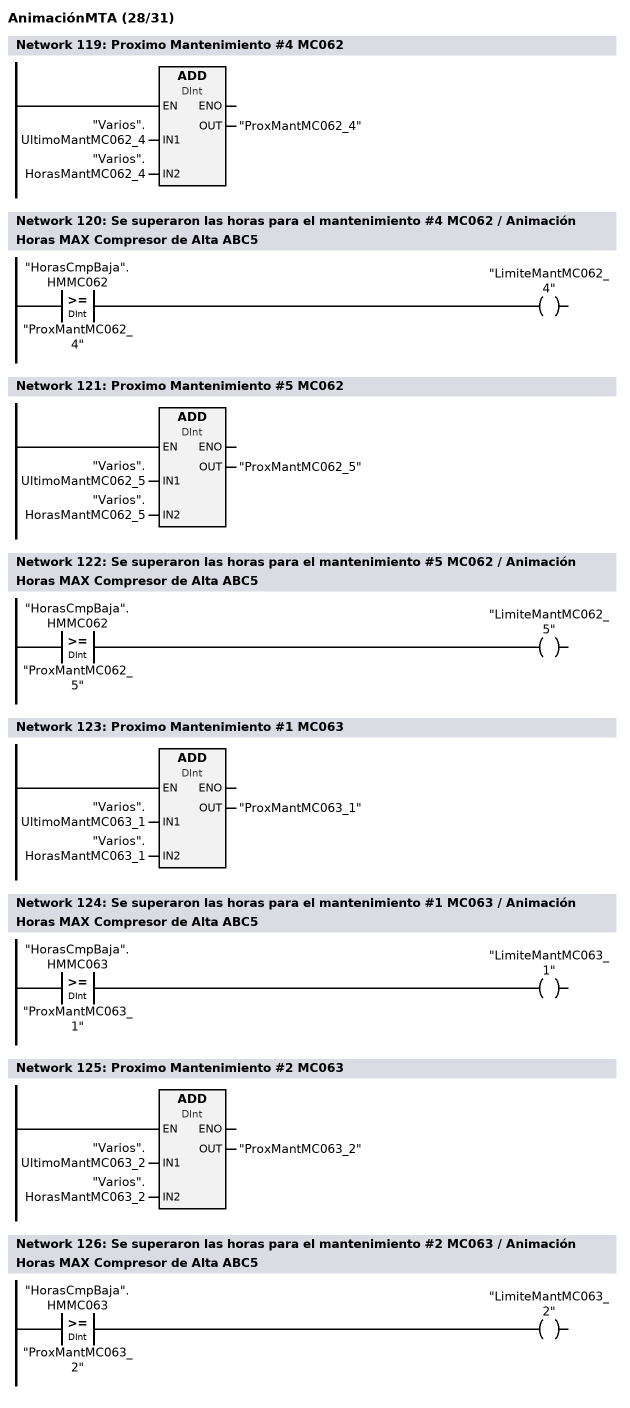
   RUNG wire#powerrail
      { S7_Templates := "SrcType := DInt"; S7_GenerateENO := "TRUE" } Add(in1 := "Varios".UltimoMantMC062_4, in2 := "Varios".HorasMantMC062_4, out => "ProxMantMC062_4")
   END_RUNG
   // the same network as SCL:
   "ProxMantMC062_4" := "Varios".UltimoMantMC062_4 + "Varios".HorasMantMC062_4;
END_REGION

REGION Network 120: Se superaron las horas para el mantenimiento #4 MC062 / Animación Horas MAX Compresor de Alta ABC5
   RUNG wire#powerrail
      { S7_Templates := "SrcType := DInt" } GE_Contact(in1 := "HorasCmpBaja".HMMC062, in2 := "ProxMantMC062_4")
      Coil( "LimiteMantMC062_4" )
   END_RUNG
   // the same network as SCL:
   "LimiteMantMC062_4" := "HorasCmpBaja".HMMC062 >= "ProxMantMC062_4";
END_REGION

REGION Network 121: Proximo Mantenimiento #5 MC062
   RUNG wire#powerrail
      { S7_Templates := "SrcType := DInt"; S7_GenerateENO := "TRUE" } Add(in1 := "Varios".UltimoMantMC062_5, in2 := "Varios".HorasMantMC062_5, out => "ProxMantMC062_5")
   END_RUNG
   // the same network as SCL:
   "ProxMantMC062_5" := "Varios".UltimoMantMC062_5 + "Varios".HorasMantMC062_5;
END_REGION

REGION Network 122: Se superaron las horas para el mantenimiento #5 MC062 / Animación Horas MAX Compresor de Alta ABC5
   RUNG wire#powerrail
      { S7_Templates := "SrcType := DInt" } GE_Contact(in1 := "HorasCmpBaja".HMMC062, in2 := "ProxMantMC062_5")
      Coil( "LimiteMantMC062_5" )
   END_RUNG
   // the same network as SCL:
   "LimiteMantMC062_5" := "HorasCmpBaja".HMMC062 >= "ProxMantMC062_5";
END_REGION

REGION Network 123: Proximo Mantenimiento #1 MC063
   RUNG wire#powerrail
      { S7_Templates := "SrcType := DInt"; S7_GenerateENO := "TRUE" } Add(in1 := "Varios".UltimoMantMC063_1, in2 := "Varios".HorasMantMC063_1, out => "ProxMantMC063_1")
   END_RUNG
   // the same network as SCL:
   "ProxMantMC063_1" := "Varios".UltimoMantMC063_1 + "Varios".HorasMantMC063_1;
END_REGION

REGION Network 124: Se superaron las horas para el mantenimiento #1 MC063 / Animación Horas MAX Compresor de Alta ABC5
   RUNG wire#powerrail
      { S7_Templates := "SrcType := DInt" } GE_Contact(in1 := "HorasCmpBaja".HMMC063, in2 := "ProxMantMC063_1")
      Coil( "LimiteMantMC063_1" )
   END_RUNG
   // the same network as SCL:
   "LimiteMantMC063_1" := "HorasCmpBaja".HMMC063 >= "ProxMantMC063_1";
END_REGION

REGION Network 125: Proximo Mantenimiento #2 MC063
   RUNG wire#powerrail
      { S7_Templates := "SrcType := DInt"; S7_GenerateENO := "TRUE" } Add(in1 := "Varios".UltimoMantMC063_2, in2 := "Varios".HorasMantMC063_2, out => "ProxMantMC063_2")
   END_RUNG
   // the same network as SCL:
   "ProxMantMC063_2" := "Varios".UltimoMantMC063_2 + "Varios".HorasMantMC063_2;
END_REGION

REGION Network 126: Se superaron las horas para el mantenimiento #2 MC063 / Animación Horas MAX Compresor de Alta ABC5
   RUNG wire#powerrail
      { S7_Templates := "SrcType := DInt" } GE_Contact(in1 := "HorasCmpBaja".HMMC063, in2 := "ProxMantMC063_2")
      Coil( "LimiteMantMC063_2" )
   END_RUNG
   // the same network as SCL:
   "LimiteMantMC063_2" := "HorasCmpBaja".HMMC063 >= "ProxMantMC063_2";
END_REGION

REGION Network 127: Proximo Mantenimiento #3 MC063
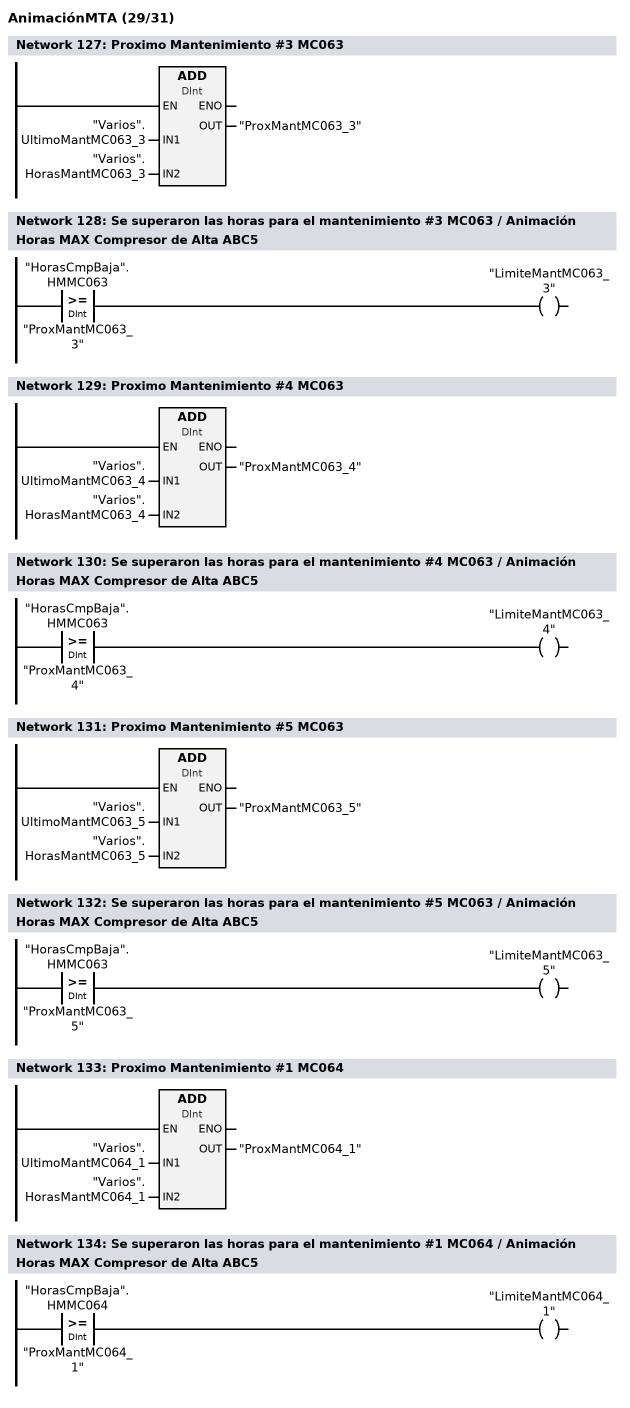
   RUNG wire#powerrail
      { S7_Templates := "SrcType := DInt"; S7_GenerateENO := "TRUE" } Add(in1 := "Varios".UltimoMantMC063_3, in2 := "Varios".HorasMantMC063_3, out => "ProxMantMC063_3")
   END_RUNG
   // the same network as SCL:
   "ProxMantMC063_3" := "Varios".UltimoMantMC063_3 + "Varios".HorasMantMC063_3;
END_REGION

REGION Network 128: Se superaron las horas para el mantenimiento #3 MC063 / Animación Horas MAX Compresor de Alta ABC5
   RUNG wire#powerrail
      { S7_Templates := "SrcType := DInt" } GE_Contact(in1 := "HorasCmpBaja".HMMC063, in2 := "ProxMantMC063_3")
      Coil( "LimiteMantMC063_3" )
   END_RUNG
   // the same network as SCL:
   "LimiteMantMC063_3" := "HorasCmpBaja".HMMC063 >= "ProxMantMC063_3";
END_REGION

REGION Network 129: Proximo Mantenimiento #4 MC063
   RUNG wire#powerrail
      { S7_Templates := "SrcType := DInt"; S7_GenerateENO := "TRUE" } Add(in1 := "Varios".UltimoMantMC063_4, in2 := "Varios".HorasMantMC063_4, out => "ProxMantMC063_4")
   END_RUNG
   // the same network as SCL:
   "ProxMantMC063_4" := "Varios".UltimoMantMC063_4 + "Varios".HorasMantMC063_4;
END_REGION

REGION Network 130: Se superaron las horas para el mantenimiento #4 MC063 / Animación Horas MAX Compresor de Alta ABC5
   RUNG wire#powerrail
      { S7_Templates := "SrcType := DInt" } GE_Contact(in1 := "HorasCmpBaja".HMMC063, in2 := "ProxMantMC063_4")
      Coil( "LimiteMantMC063_4" )
   END_RUNG
   // the same network as SCL:
   "LimiteMantMC063_4" := "HorasCmpBaja".HMMC063 >= "ProxMantMC063_4";
END_REGION

REGION Network 131: Proximo Mantenimiento #5 MC063
   RUNG wire#powerrail
      { S7_Templates := "SrcType := DInt"; S7_GenerateENO := "TRUE" } Add(in1 := "Varios".UltimoMantMC063_5, in2 := "Varios".HorasMantMC063_5, out => "ProxMantMC063_5")
   END_RUNG
   // the same network as SCL:
   "ProxMantMC063_5" := "Varios".UltimoMantMC063_5 + "Varios".HorasMantMC063_5;
END_REGION

REGION Network 132: Se superaron las horas para el mantenimiento #5 MC063 / Animación Horas MAX Compresor de Alta ABC5
   RUNG wire#powerrail
      { S7_Templates := "SrcType := DInt" } GE_Contact(in1 := "HorasCmpBaja".HMMC063, in2 := "ProxMantMC063_5")
      Coil( "LimiteMantMC063_5" )
   END_RUNG
   // the same network as SCL:
   "LimiteMantMC063_5" := "HorasCmpBaja".HMMC063 >= "ProxMantMC063_5";
END_REGION

REGION Network 133: Proximo Mantenimiento #1 MC064
   RUNG wire#powerrail
      { S7_Templates := "SrcType := DInt"; S7_GenerateENO := "TRUE" } Add(in1 := "Varios".UltimoMantMC064_1, in2 := "Varios".HorasMantMC064_1, out => "ProxMantMC064_1")
   END_RUNG
   // the same network as SCL:
   "ProxMantMC064_1" := "Varios".UltimoMantMC064_1 + "Varios".HorasMantMC064_1;
END_REGION

REGION Network 134: Se superaron las horas para el mantenimiento #1 MC064 / Animación Horas MAX Compresor de Alta ABC5
   RUNG wire#powerrail
      { S7_Templates := "SrcType := DInt" } GE_Contact(in1 := "HorasCmpBaja".HMMC064, in2 := "ProxMantMC064_1")
      Coil( "LimiteMantMC064_1" )
   END_RUNG
   // the same network as SCL:
   "LimiteMantMC064_1" := "HorasCmpBaja".HMMC064 >= "ProxMantMC064_1";
END_REGION

REGION Network 135: Proximo Mantenimiento #2 MC064
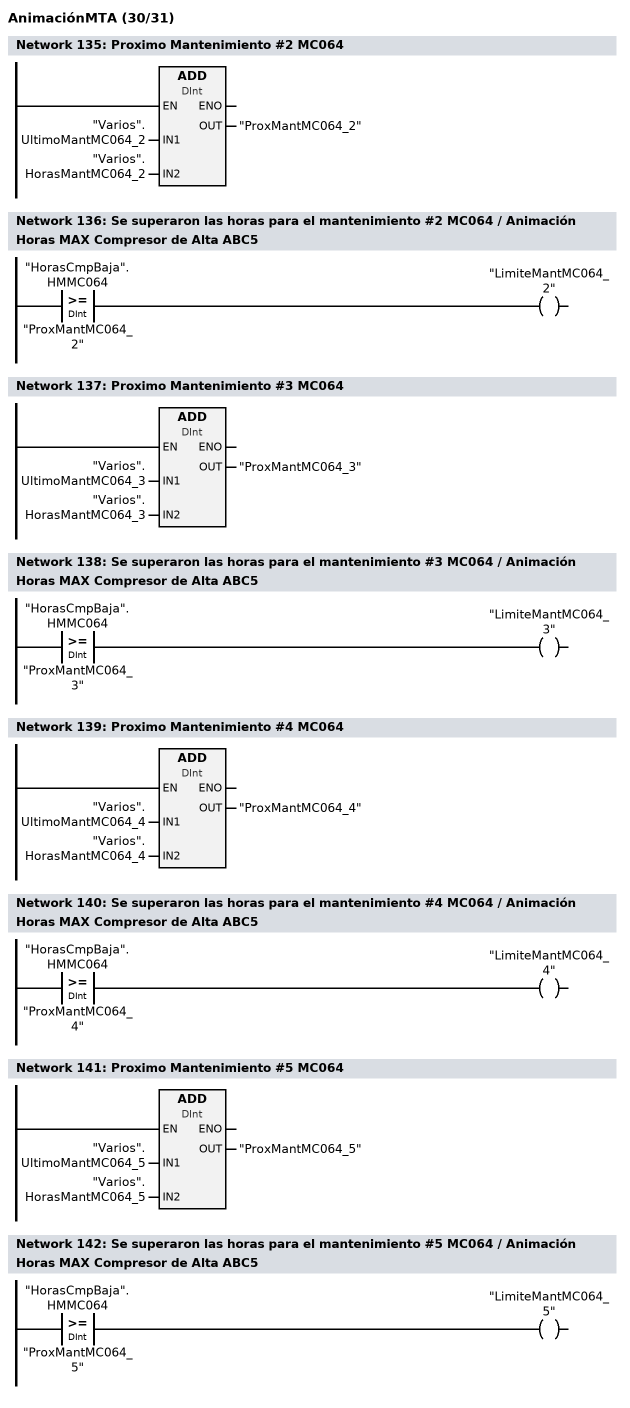
   RUNG wire#powerrail
      { S7_Templates := "SrcType := DInt"; S7_GenerateENO := "TRUE" } Add(in1 := "Varios".UltimoMantMC064_2, in2 := "Varios".HorasMantMC064_2, out => "ProxMantMC064_2")
   END_RUNG
   // the same network as SCL:
   "ProxMantMC064_2" := "Varios".UltimoMantMC064_2 + "Varios".HorasMantMC064_2;
END_REGION

REGION Network 136: Se superaron las horas para el mantenimiento #2 MC064 / Animación Horas MAX Compresor de Alta ABC5
   RUNG wire#powerrail
      { S7_Templates := "SrcType := DInt" } GE_Contact(in1 := "HorasCmpBaja".HMMC064, in2 := "ProxMantMC064_2")
      Coil( "LimiteMantMC064_2" )
   END_RUNG
   // the same network as SCL:
   "LimiteMantMC064_2" := "HorasCmpBaja".HMMC064 >= "ProxMantMC064_2";
END_REGION

REGION Network 137: Proximo Mantenimiento #3 MC064
   RUNG wire#powerrail
      { S7_Templates := "SrcType := DInt"; S7_GenerateENO := "TRUE" } Add(in1 := "Varios".UltimoMantMC064_3, in2 := "Varios".HorasMantMC064_3, out => "ProxMantMC064_3")
   END_RUNG
   // the same network as SCL:
   "ProxMantMC064_3" := "Varios".UltimoMantMC064_3 + "Varios".HorasMantMC064_3;
END_REGION

REGION Network 138: Se superaron las horas para el mantenimiento #3 MC064 / Animación Horas MAX Compresor de Alta ABC5
   RUNG wire#powerrail
      { S7_Templates := "SrcType := DInt" } GE_Contact(in1 := "HorasCmpBaja".HMMC064, in2 := "ProxMantMC064_3")
      Coil( "LimiteMantMC064_3" )
   END_RUNG
   // the same network as SCL:
   "LimiteMantMC064_3" := "HorasCmpBaja".HMMC064 >= "ProxMantMC064_3";
END_REGION

REGION Network 139: Proximo Mantenimiento #4 MC064
   RUNG wire#powerrail
      { S7_Templates := "SrcType := DInt"; S7_GenerateENO := "TRUE" } Add(in1 := "Varios".UltimoMantMC064_4, in2 := "Varios".HorasMantMC064_4, out => "ProxMantMC064_4")
   END_RUNG
   // the same network as SCL:
   "ProxMantMC064_4" := "Varios".UltimoMantMC064_4 + "Varios".HorasMantMC064_4;
END_REGION

REGION Network 140: Se superaron las horas para el mantenimiento #4 MC064 / Animación Horas MAX Compresor de Alta ABC5
   RUNG wire#powerrail
      { S7_Templates := "SrcType := DInt" } GE_Contact(in1 := "HorasCmpBaja".HMMC064, in2 := "ProxMantMC064_4")
      Coil( "LimiteMantMC064_4" )
   END_RUNG
   // the same network as SCL:
   "LimiteMantMC064_4" := "HorasCmpBaja".HMMC064 >= "ProxMantMC064_4";
END_REGION

REGION Network 141: Proximo Mantenimiento #5 MC064
   RUNG wire#powerrail
      { S7_Templates := "SrcType := DInt"; S7_GenerateENO := "TRUE" } Add(in1 := "Varios".UltimoMantMC064_5, in2 := "Varios".HorasMantMC064_5, out => "ProxMantMC064_5")
   END_RUNG
   // the same network as SCL:
   "ProxMantMC064_5" := "Varios".UltimoMantMC064_5 + "Varios".HorasMantMC064_5;
END_REGION

REGION Network 142: Se superaron las horas para el mantenimiento #5 MC064 / Animación Horas MAX Compresor de Alta ABC5
   RUNG wire#powerrail
      { S7_Templates := "SrcType := DInt" } GE_Contact(in1 := "HorasCmpBaja".HMMC064, in2 := "ProxMantMC064_5")
      Coil( "LimiteMantMC064_5" )
   END_RUNG
   // the same network as SCL:
   "LimiteMantMC064_5" := "HorasCmpBaja".HMMC064 >= "ProxMantMC064_5";
END_REGION

REGION Network 143: Próximo Mantenimento Booster 1
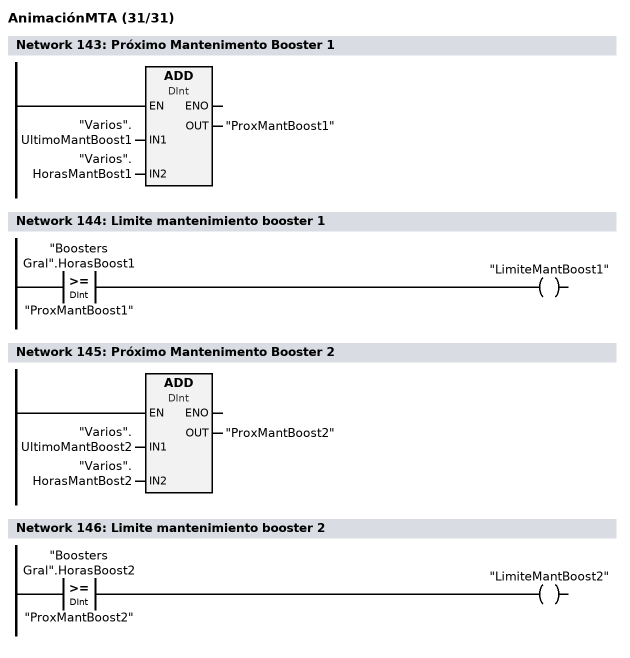
   RUNG wire#powerrail
      { S7_Templates := "SrcType := DInt"; S7_GenerateENO := "TRUE" } Add(in1 := "Varios".UltimoMantBoost1, in2 := "Varios".HorasMantBost1, out => "ProxMantBoost1")
   END_RUNG
   // the same network as SCL:
   "ProxMantBoost1" := "Varios".UltimoMantBoost1 + "Varios".HorasMantBost1;
END_REGION

REGION Network 144: Limite mantenimiento booster 1
   RUNG wire#powerrail
      { S7_Templates := "SrcType := DInt" } GE_Contact(in1 := "Boosters Gral".HorasBoost1, in2 := "ProxMantBoost1")
      Coil( "LimiteMantBoost1" )
   END_RUNG
   // the same network as SCL:
   "LimiteMantBoost1" := "Boosters Gral".HorasBoost1 >= "ProxMantBoost1";
END_REGION

REGION Network 145: Próximo Mantenimento Booster 2
   RUNG wire#powerrail
      { S7_Templates := "SrcType := DInt"; S7_GenerateENO := "TRUE" } Add(in1 := "Varios".UltimoMantBoost2, in2 := "Varios".HorasMantBost2, out => "ProxMantBoost2")
   END_RUNG
   // the same network as SCL:
   "ProxMantBoost2" := "Varios".UltimoMantBoost2 + "Varios".HorasMantBost2;
END_REGION

REGION Network 146: Limite mantenimiento booster 2
   RUNG wire#powerrail
      { S7_Templates := "SrcType := DInt" } GE_Contact(in1 := "Boosters Gral".HorasBoost2, in2 := "ProxMantBoost2")
      Coil( "LimiteMantBoost2" )
   END_RUNG
   // the same network as SCL:
   "LimiteMantBoost2" := "Boosters Gral".HorasBoost2 >= "ProxMantBoost2";
END_REGION
END_FUNCTION

FUNCTION "Motores-PanelMTA" : Void   // FC3, LAD
{ S7_Optimized_Access := 'FALSE' }
VERSION : 0.1
BEGIN

REGION Network 1: Comandos desde Panel para MP010 - Bomba Principal Ch. Soplado
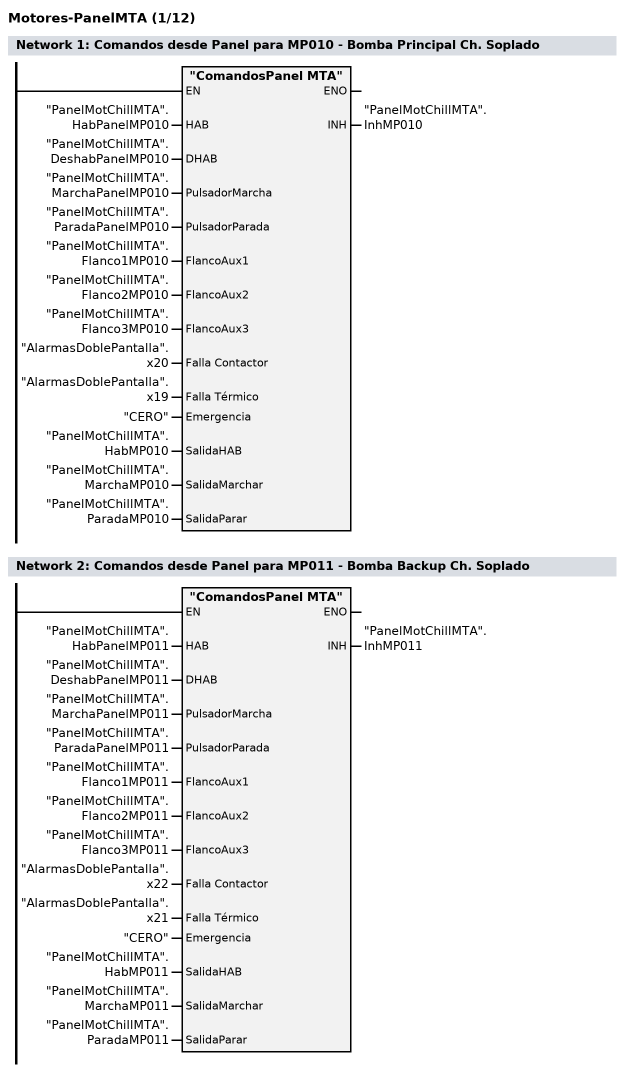
   RUNG wire#powerrail
      "ComandosPanel MTA"(HAB := "PanelMotChillMTA".HabPanelMP010, DHAB := "PanelMotChillMTA".DeshabPanelMP010, PulsadorMarcha := "PanelMotChillMTA".MarchaPanelMP010, PulsadorParada := "PanelMotChillMTA".ParadaPanelMP010, FlancoAux1 := "PanelMotChillMTA".Flanco1MP010, FlancoAux2 := "PanelMotChillMTA".Flanco2MP010, FlancoAux3 := "PanelMotChillMTA".Flanco3MP010, "Falla Contactor" := "AlarmasDoblePantalla".x20, "Falla Térmico" := "AlarmasDoblePantalla".x19, Emergencia := "CERO", INH => "PanelMotChillMTA".InhMP010, SalidaHAB := "PanelMotChillMTA".HabMP010, SalidaMarchar := "PanelMotChillMTA".MarchaMP010, SalidaParar := "PanelMotChillMTA".ParadaMP010)
   END_RUNG
   // the same network as SCL:
   "ComandosPanel MTA"(HAB := "PanelMotChillMTA".HabPanelMP010,
                       DHAB := "PanelMotChillMTA".DeshabPanelMP010,
                       PulsadorMarcha := "PanelMotChillMTA".MarchaPanelMP010,
                       PulsadorParada := "PanelMotChillMTA".ParadaPanelMP010,
                       FlancoAux1 := "PanelMotChillMTA".Flanco1MP010,
                       FlancoAux2 := "PanelMotChillMTA".Flanco2MP010,
                       FlancoAux3 := "PanelMotChillMTA".Flanco3MP010,
                       "Falla Contactor" := "AlarmasDoblePantalla".x20,
                       "Falla Térmico" := "AlarmasDoblePantalla".x19,
                       Emergencia := "CERO",
                       SalidaHAB := "PanelMotChillMTA".HabMP010,
                       SalidaMarchar := "PanelMotChillMTA".MarchaMP010,
                       SalidaParar := "PanelMotChillMTA".ParadaMP010,
                       INH => "PanelMotChillMTA".InhMP010);
END_REGION

REGION Network 2: Comandos desde Panel para MP011 - Bomba Backup Ch. Soplado
   RUNG wire#powerrail
      "ComandosPanel MTA"(HAB := "PanelMotChillMTA".HabPanelMP011, DHAB := "PanelMotChillMTA".DeshabPanelMP011, PulsadorMarcha := "PanelMotChillMTA".MarchaPanelMP011, PulsadorParada := "PanelMotChillMTA".ParadaPanelMP011, FlancoAux1 := "PanelMotChillMTA".Flanco1MP011, FlancoAux2 := "PanelMotChillMTA".Flanco2MP011, FlancoAux3 := "PanelMotChillMTA".Flanco3MP011, "Falla Contactor" := "AlarmasDoblePantalla".x22, "Falla Térmico" := "AlarmasDoblePantalla".x21, Emergencia := "CERO", INH => "PanelMotChillMTA".InhMP011, SalidaHAB := "PanelMotChillMTA".HabMP011, SalidaMarchar := "PanelMotChillMTA".MarchaMP011, SalidaParar := "PanelMotChillMTA".ParadaMP011)
   END_RUNG
   // the same network as SCL:
   "ComandosPanel MTA"(HAB := "PanelMotChillMTA".HabPanelMP011,
                       DHAB := "PanelMotChillMTA".DeshabPanelMP011,
                       PulsadorMarcha := "PanelMotChillMTA".MarchaPanelMP011,
                       PulsadorParada := "PanelMotChillMTA".ParadaPanelMP011,
                       FlancoAux1 := "PanelMotChillMTA".Flanco1MP011,
                       FlancoAux2 := "PanelMotChillMTA".Flanco2MP011,
                       FlancoAux3 := "PanelMotChillMTA".Flanco3MP011,
                       "Falla Contactor" := "AlarmasDoblePantalla".x22,
                       "Falla Térmico" := "AlarmasDoblePantalla".x21,
                       Emergencia := "CERO",
                       SalidaHAB := "PanelMotChillMTA".HabMP011,
                       SalidaMarchar := "PanelMotChillMTA".MarchaMP011,
                       SalidaParar := "PanelMotChillMTA".ParadaMP011,
                       INH => "PanelMotChillMTA".InhMP011);
END_REGION

REGION Network 3: Comandos desde Panel para MP012 - Bomba Principal Ch. Envasado
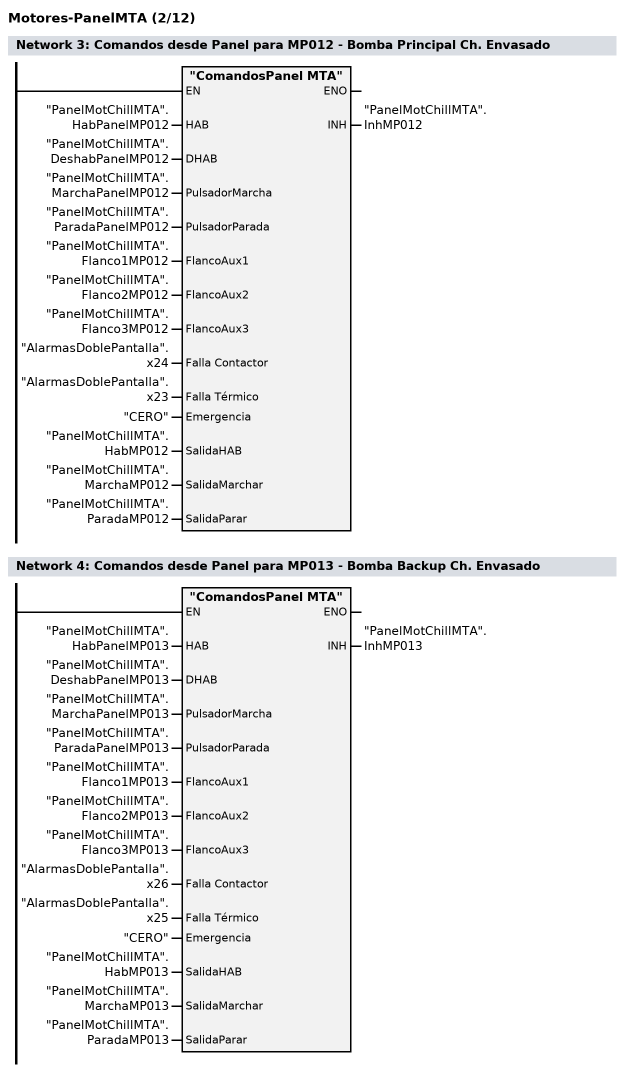
   RUNG wire#powerrail
      "ComandosPanel MTA"(HAB := "PanelMotChillMTA".HabPanelMP012, DHAB := "PanelMotChillMTA".DeshabPanelMP012, PulsadorMarcha := "PanelMotChillMTA".MarchaPanelMP012, PulsadorParada := "PanelMotChillMTA".ParadaPanelMP012, FlancoAux1 := "PanelMotChillMTA".Flanco1MP012, FlancoAux2 := "PanelMotChillMTA".Flanco2MP012, FlancoAux3 := "PanelMotChillMTA".Flanco3MP012, "Falla Contactor" := "AlarmasDoblePantalla".x24, "Falla Térmico" := "AlarmasDoblePantalla".x23, Emergencia := "CERO", INH => "PanelMotChillMTA".InhMP012, SalidaHAB := "PanelMotChillMTA".HabMP012, SalidaMarchar := "PanelMotChillMTA".MarchaMP012, SalidaParar := "PanelMotChillMTA".ParadaMP012)
   END_RUNG
   // the same network as SCL:
   "ComandosPanel MTA"(HAB := "PanelMotChillMTA".HabPanelMP012,
                       DHAB := "PanelMotChillMTA".DeshabPanelMP012,
                       PulsadorMarcha := "PanelMotChillMTA".MarchaPanelMP012,
                       PulsadorParada := "PanelMotChillMTA".ParadaPanelMP012,
                       FlancoAux1 := "PanelMotChillMTA".Flanco1MP012,
                       FlancoAux2 := "PanelMotChillMTA".Flanco2MP012,
                       FlancoAux3 := "PanelMotChillMTA".Flanco3MP012,
                       "Falla Contactor" := "AlarmasDoblePantalla".x24,
                       "Falla Térmico" := "AlarmasDoblePantalla".x23,
                       Emergencia := "CERO",
                       SalidaHAB := "PanelMotChillMTA".HabMP012,
                       SalidaMarchar := "PanelMotChillMTA".MarchaMP012,
                       SalidaParar := "PanelMotChillMTA".ParadaMP012,
                       INH => "PanelMotChillMTA".InhMP012);
END_REGION

REGION Network 4: Comandos desde Panel para MP013 - Bomba Backup Ch. Envasado
   RUNG wire#powerrail
      "ComandosPanel MTA"(HAB := "PanelMotChillMTA".HabPanelMP013, DHAB := "PanelMotChillMTA".DeshabPanelMP013, PulsadorMarcha := "PanelMotChillMTA".MarchaPanelMP013, PulsadorParada := "PanelMotChillMTA".ParadaPanelMP013, FlancoAux1 := "PanelMotChillMTA".Flanco1MP013, FlancoAux2 := "PanelMotChillMTA".Flanco2MP013, FlancoAux3 := "PanelMotChillMTA".Flanco3MP013, "Falla Contactor" := "AlarmasDoblePantalla".x26, "Falla Térmico" := "AlarmasDoblePantalla".x25, Emergencia := "CERO", INH => "PanelMotChillMTA".InhMP013, SalidaHAB := "PanelMotChillMTA".HabMP013, SalidaMarchar := "PanelMotChillMTA".MarchaMP013, SalidaParar := "PanelMotChillMTA".ParadaMP013)
   END_RUNG
   // the same network as SCL:
   "ComandosPanel MTA"(HAB := "PanelMotChillMTA".HabPanelMP013,
                       DHAB := "PanelMotChillMTA".DeshabPanelMP013,
                       PulsadorMarcha := "PanelMotChillMTA".MarchaPanelMP013,
                       PulsadorParada := "PanelMotChillMTA".ParadaPanelMP013,
                       FlancoAux1 := "PanelMotChillMTA".Flanco1MP013,
                       FlancoAux2 := "PanelMotChillMTA".Flanco2MP013,
                       FlancoAux3 := "PanelMotChillMTA".Flanco3MP013,
                       "Falla Contactor" := "AlarmasDoblePantalla".x26,
                       "Falla Térmico" := "AlarmasDoblePantalla".x25,
                       Emergencia := "CERO",
                       SalidaHAB := "PanelMotChillMTA".HabMP013,
                       SalidaMarchar := "PanelMotChillMTA".MarchaMP013,
                       SalidaParar := "PanelMotChillMTA".ParadaMP013,
                       INH => "PanelMotChillMTA".InhMP013);
END_REGION

REGION Network 5: Comandos desde Panel para MP018 - Bomba 1 Torres de enfriamiento Chillers
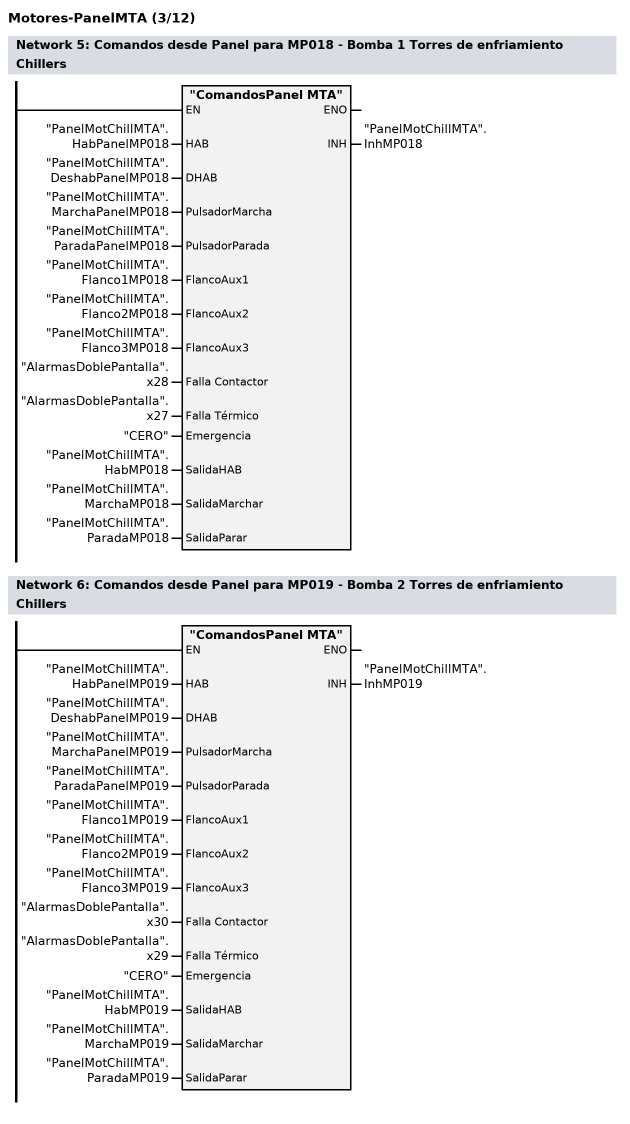
   RUNG wire#powerrail
      "ComandosPanel MTA"(HAB := "PanelMotChillMTA".HabPanelMP018, DHAB := "PanelMotChillMTA".DeshabPanelMP018, PulsadorMarcha := "PanelMotChillMTA".MarchaPanelMP018, PulsadorParada := "PanelMotChillMTA".ParadaPanelMP018, FlancoAux1 := "PanelMotChillMTA".Flanco1MP018, FlancoAux2 := "PanelMotChillMTA".Flanco2MP018, FlancoAux3 := "PanelMotChillMTA".Flanco3MP018, "Falla Contactor" := "AlarmasDoblePantalla".x28, "Falla Térmico" := "AlarmasDoblePantalla".x27, Emergencia := "CERO", SalidaHAB := "PanelMotChillMTA".HabMP018, SalidaMarchar := "PanelMotChillMTA".MarchaMP018, SalidaParar := "PanelMotChillMTA".ParadaMP018, INH => "PanelMotChillMTA".InhMP018)
   END_RUNG
   // the same network as SCL:
   "ComandosPanel MTA"(HAB := "PanelMotChillMTA".HabPanelMP018,
                       DHAB := "PanelMotChillMTA".DeshabPanelMP018,
                       PulsadorMarcha := "PanelMotChillMTA".MarchaPanelMP018,
                       PulsadorParada := "PanelMotChillMTA".ParadaPanelMP018,
                       FlancoAux1 := "PanelMotChillMTA".Flanco1MP018,
                       FlancoAux2 := "PanelMotChillMTA".Flanco2MP018,
                       FlancoAux3 := "PanelMotChillMTA".Flanco3MP018,
                       "Falla Contactor" := "AlarmasDoblePantalla".x28,
                       "Falla Térmico" := "AlarmasDoblePantalla".x27,
                       Emergencia := "CERO",
                       SalidaHAB := "PanelMotChillMTA".HabMP018,
                       SalidaMarchar := "PanelMotChillMTA".MarchaMP018,
                       SalidaParar := "PanelMotChillMTA".ParadaMP018,
                       INH => "PanelMotChillMTA".InhMP018);
END_REGION

REGION Network 6: Comandos desde Panel para MP019 - Bomba 2 Torres de enfriamiento Chillers
   RUNG wire#powerrail
      "ComandosPanel MTA"(HAB := "PanelMotChillMTA".HabPanelMP019, DHAB := "PanelMotChillMTA".DeshabPanelMP019, PulsadorMarcha := "PanelMotChillMTA".MarchaPanelMP019, PulsadorParada := "PanelMotChillMTA".ParadaPanelMP019, FlancoAux1 := "PanelMotChillMTA".Flanco1MP019, FlancoAux2 := "PanelMotChillMTA".Flanco2MP019, FlancoAux3 := "PanelMotChillMTA".Flanco3MP019, "Falla Contactor" := "AlarmasDoblePantalla".x30, "Falla Térmico" := "AlarmasDoblePantalla".x29, Emergencia := "CERO", SalidaHAB := "PanelMotChillMTA".HabMP019, SalidaMarchar := "PanelMotChillMTA".MarchaMP019, SalidaParar := "PanelMotChillMTA".ParadaMP019, INH => "PanelMotChillMTA".InhMP019)
   END_RUNG
   // the same network as SCL:
   "ComandosPanel MTA"(HAB := "PanelMotChillMTA".HabPanelMP019,
                       DHAB := "PanelMotChillMTA".DeshabPanelMP019,
                       PulsadorMarcha := "PanelMotChillMTA".MarchaPanelMP019,
                       PulsadorParada := "PanelMotChillMTA".ParadaPanelMP019,
                       FlancoAux1 := "PanelMotChillMTA".Flanco1MP019,
                       FlancoAux2 := "PanelMotChillMTA".Flanco2MP019,
                       FlancoAux3 := "PanelMotChillMTA".Flanco3MP019,
                       "Falla Contactor" := "AlarmasDoblePantalla".x30,
                       "Falla Térmico" := "AlarmasDoblePantalla".x29,
                       Emergencia := "CERO",
                       SalidaHAB := "PanelMotChillMTA".HabMP019,
                       SalidaMarchar := "PanelMotChillMTA".MarchaMP019,
                       SalidaParar := "PanelMotChillMTA".ParadaMP019,
                       INH => "PanelMotChillMTA".InhMP019);
END_REGION

REGION Network 7: Comandos desde Panel para MT007 - Bomba Soplado L1
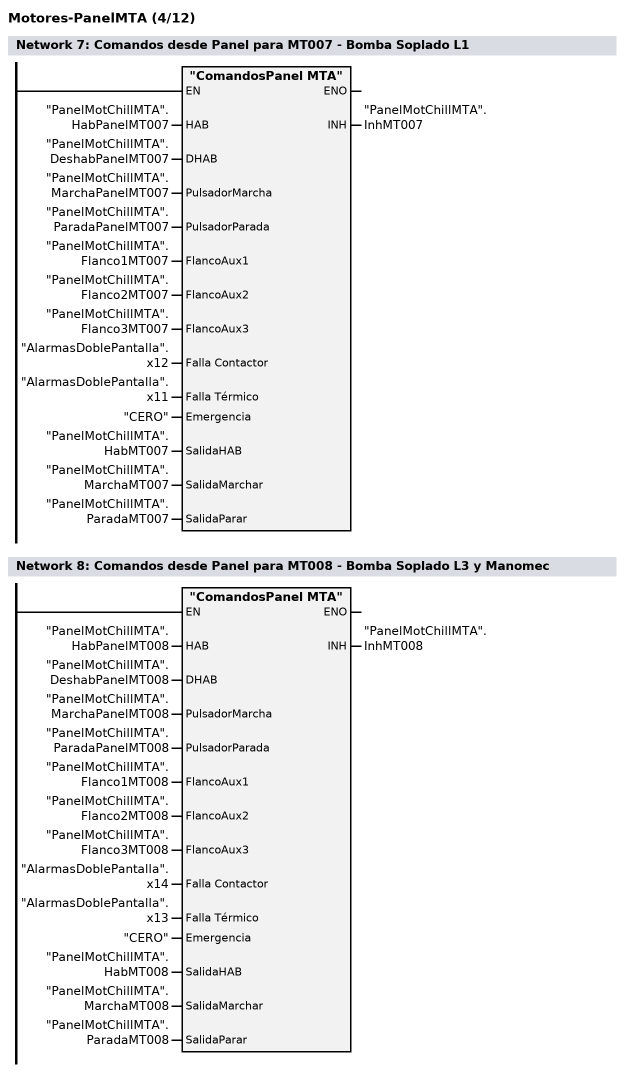
   RUNG wire#powerrail
      "ComandosPanel MTA"(HAB := "PanelMotChillMTA".HabPanelMT007, DHAB := "PanelMotChillMTA".DeshabPanelMT007, PulsadorMarcha := "PanelMotChillMTA".MarchaPanelMT007, PulsadorParada := "PanelMotChillMTA".ParadaPanelMT007, FlancoAux1 := "PanelMotChillMTA".Flanco1MT007, FlancoAux2 := "PanelMotChillMTA".Flanco2MT007, FlancoAux3 := "PanelMotChillMTA".Flanco3MT007, "Falla Contactor" := "AlarmasDoblePantalla".x12, "Falla Térmico" := "AlarmasDoblePantalla".x11, Emergencia := "CERO", INH => "PanelMotChillMTA".InhMT007, SalidaHAB := "PanelMotChillMTA".HabMT007, SalidaMarchar := "PanelMotChillMTA".MarchaMT007, SalidaParar := "PanelMotChillMTA".ParadaMT007)
   END_RUNG
   // the same network as SCL:
   "ComandosPanel MTA"(HAB := "PanelMotChillMTA".HabPanelMT007,
                       DHAB := "PanelMotChillMTA".DeshabPanelMT007,
                       PulsadorMarcha := "PanelMotChillMTA".MarchaPanelMT007,
                       PulsadorParada := "PanelMotChillMTA".ParadaPanelMT007,
                       FlancoAux1 := "PanelMotChillMTA".Flanco1MT007,
                       FlancoAux2 := "PanelMotChillMTA".Flanco2MT007,
                       FlancoAux3 := "PanelMotChillMTA".Flanco3MT007,
                       "Falla Contactor" := "AlarmasDoblePantalla".x12,
                       "Falla Térmico" := "AlarmasDoblePantalla".x11,
                       Emergencia := "CERO",
                       SalidaHAB := "PanelMotChillMTA".HabMT007,
                       SalidaMarchar := "PanelMotChillMTA".MarchaMT007,
                       SalidaParar := "PanelMotChillMTA".ParadaMT007,
                       INH => "PanelMotChillMTA".InhMT007);
END_REGION

REGION Network 8: Comandos desde Panel para MT008 - Bomba Soplado L3 y Manomec
   RUNG wire#powerrail
      "ComandosPanel MTA"(HAB := "PanelMotChillMTA".HabPanelMT008, DHAB := "PanelMotChillMTA".DeshabPanelMT008, PulsadorMarcha := "PanelMotChillMTA".MarchaPanelMT008, PulsadorParada := "PanelMotChillMTA".ParadaPanelMT008, FlancoAux1 := "PanelMotChillMTA".Flanco1MT008, FlancoAux2 := "PanelMotChillMTA".Flanco2MT008, FlancoAux3 := "PanelMotChillMTA".Flanco3MT008, "Falla Contactor" := "AlarmasDoblePantalla".x14, "Falla Térmico" := "AlarmasDoblePantalla".x13, Emergencia := "CERO", INH => "PanelMotChillMTA".InhMT008, SalidaHAB := "PanelMotChillMTA".HabMT008, SalidaMarchar := "PanelMotChillMTA".MarchaMT008, SalidaParar := "PanelMotChillMTA".ParadaMT008)
   END_RUNG
   // the same network as SCL:
   "ComandosPanel MTA"(HAB := "PanelMotChillMTA".HabPanelMT008,
                       DHAB := "PanelMotChillMTA".DeshabPanelMT008,
                       PulsadorMarcha := "PanelMotChillMTA".MarchaPanelMT008,
                       PulsadorParada := "PanelMotChillMTA".ParadaPanelMT008,
                       FlancoAux1 := "PanelMotChillMTA".Flanco1MT008,
                       FlancoAux2 := "PanelMotChillMTA".Flanco2MT008,
                       FlancoAux3 := "PanelMotChillMTA".Flanco3MT008,
                       "Falla Contactor" := "AlarmasDoblePantalla".x14,
                       "Falla Térmico" := "AlarmasDoblePantalla".x13,
                       Emergencia := "CERO",
                       SalidaHAB := "PanelMotChillMTA".HabMT008,
                       SalidaMarchar := "PanelMotChillMTA".MarchaMT008,
                       SalidaParar := "PanelMotChillMTA".ParadaMT008,
                       INH => "PanelMotChillMTA".InhMT008);
END_REGION

REGION Network 9: Comandos desde Panel para MT009 - Bomba Int. L3 y L5
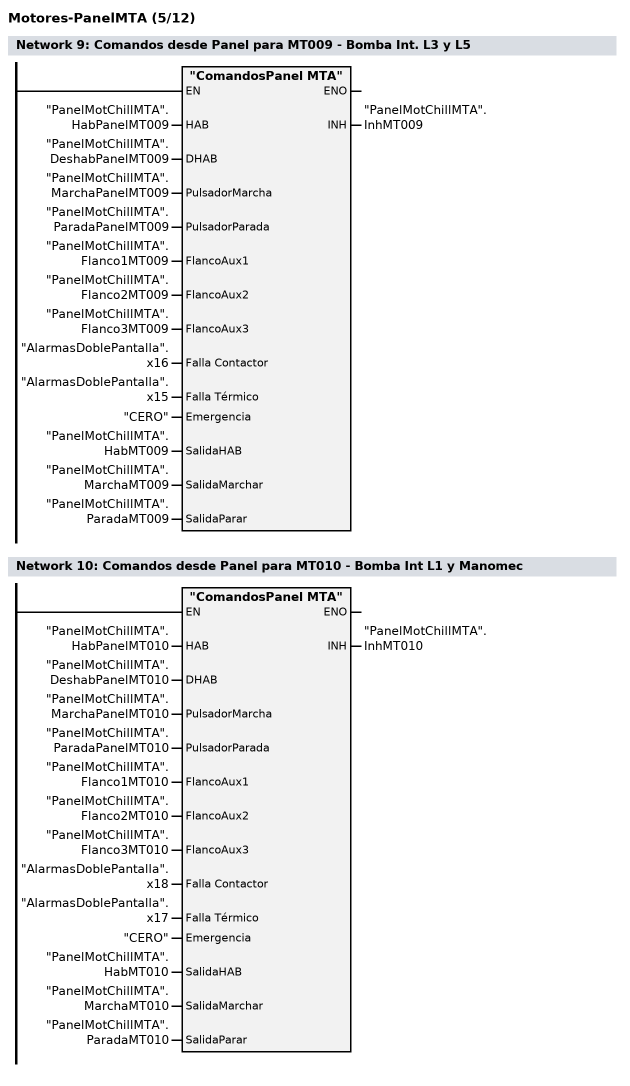
   RUNG wire#powerrail
      "ComandosPanel MTA"(HAB := "PanelMotChillMTA".HabPanelMT009, DHAB := "PanelMotChillMTA".DeshabPanelMT009, PulsadorMarcha := "PanelMotChillMTA".MarchaPanelMT009, PulsadorParada := "PanelMotChillMTA".ParadaPanelMT009, FlancoAux1 := "PanelMotChillMTA".Flanco1MT009, FlancoAux2 := "PanelMotChillMTA".Flanco2MT009, FlancoAux3 := "PanelMotChillMTA".Flanco3MT009, "Falla Contactor" := "AlarmasDoblePantalla".x16, "Falla Térmico" := "AlarmasDoblePantalla".x15, Emergencia := "CERO", INH => "PanelMotChillMTA".InhMT009, SalidaHAB := "PanelMotChillMTA".HabMT009, SalidaMarchar := "PanelMotChillMTA".MarchaMT009, SalidaParar := "PanelMotChillMTA".ParadaMT009)
   END_RUNG
   // the same network as SCL:
   "ComandosPanel MTA"(HAB := "PanelMotChillMTA".HabPanelMT009,
                       DHAB := "PanelMotChillMTA".DeshabPanelMT009,
                       PulsadorMarcha := "PanelMotChillMTA".MarchaPanelMT009,
                       PulsadorParada := "PanelMotChillMTA".ParadaPanelMT009,
                       FlancoAux1 := "PanelMotChillMTA".Flanco1MT009,
                       FlancoAux2 := "PanelMotChillMTA".Flanco2MT009,
                       FlancoAux3 := "PanelMotChillMTA".Flanco3MT009,
                       "Falla Contactor" := "AlarmasDoblePantalla".x16,
                       "Falla Térmico" := "AlarmasDoblePantalla".x15,
                       Emergencia := "CERO",
                       SalidaHAB := "PanelMotChillMTA".HabMT009,
                       SalidaMarchar := "PanelMotChillMTA".MarchaMT009,
                       SalidaParar := "PanelMotChillMTA".ParadaMT009,
                       INH => "PanelMotChillMTA".InhMT009);
END_REGION

REGION Network 10: Comandos desde Panel para MT010 - Bomba Int L1 y Manomec
   RUNG wire#powerrail
      "ComandosPanel MTA"(HAB := "PanelMotChillMTA".HabPanelMT010, DHAB := "PanelMotChillMTA".DeshabPanelMT010, PulsadorMarcha := "PanelMotChillMTA".MarchaPanelMT010, PulsadorParada := "PanelMotChillMTA".ParadaPanelMT010, FlancoAux1 := "PanelMotChillMTA".Flanco1MT010, FlancoAux2 := "PanelMotChillMTA".Flanco2MT010, FlancoAux3 := "PanelMotChillMTA".Flanco3MT010, "Falla Contactor" := "AlarmasDoblePantalla".x18, "Falla Térmico" := "AlarmasDoblePantalla".x17, Emergencia := "CERO", INH => "PanelMotChillMTA".InhMT010, SalidaHAB := "PanelMotChillMTA".HabMT010, SalidaMarchar := "PanelMotChillMTA".MarchaMT010, SalidaParar := "PanelMotChillMTA".ParadaMT010)
   END_RUNG
   // the same network as SCL:
   "ComandosPanel MTA"(HAB := "PanelMotChillMTA".HabPanelMT010,
                       DHAB := "PanelMotChillMTA".DeshabPanelMT010,
                       PulsadorMarcha := "PanelMotChillMTA".MarchaPanelMT010,
                       PulsadorParada := "PanelMotChillMTA".ParadaPanelMT010,
                       FlancoAux1 := "PanelMotChillMTA".Flanco1MT010,
                       FlancoAux2 := "PanelMotChillMTA".Flanco2MT010,
                       FlancoAux3 := "PanelMotChillMTA".Flanco3MT010,
                       "Falla Contactor" := "AlarmasDoblePantalla".x18,
                       "Falla Térmico" := "AlarmasDoblePantalla".x17,
                       Emergencia := "CERO",
                       SalidaHAB := "PanelMotChillMTA".HabMT010,
                       SalidaMarchar := "PanelMotChillMTA".MarchaMT010,
                       SalidaParar := "PanelMotChillMTA".ParadaMT010,
                       INH => "PanelMotChillMTA".InhMT010);
END_REGION

REGION Network 11: Comandos desde Panel para V001 - Ventilador 1 Torres de enfriamiento Chillers
